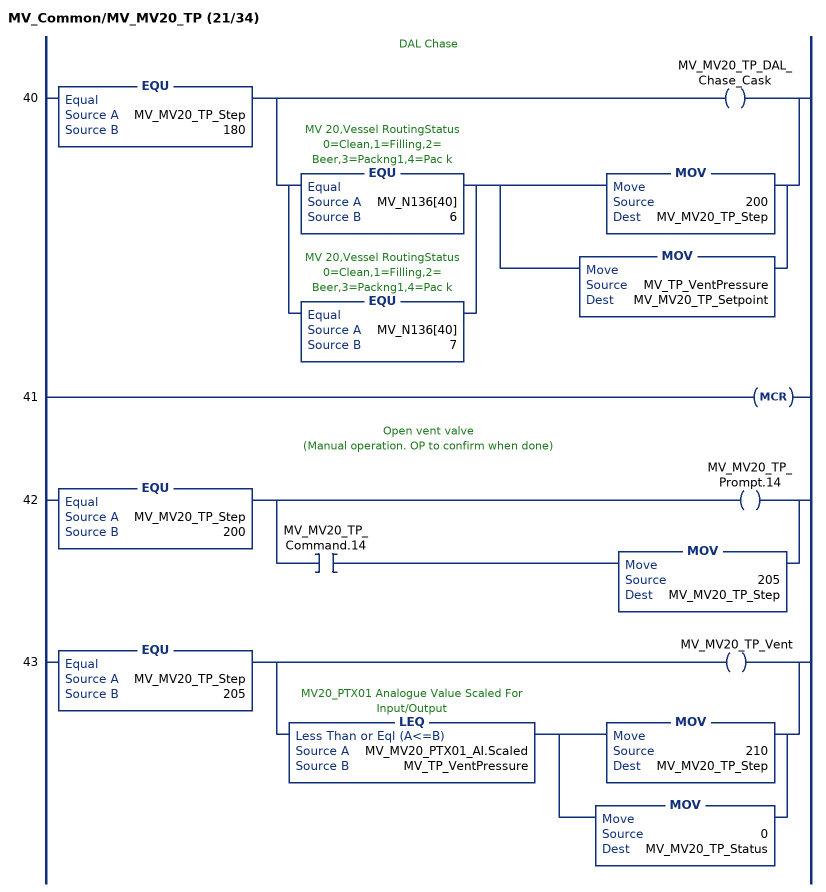
   // DAL Chase
   40: EQU(MV_MV20_TP_Step,180)[OTE(MV_MV20_TP_DAL_Chase_Cask) ,[EQU(MV_N136[40],6) ,EQU(MV_N136[40],7) ] [MOV(200,MV_MV20_TP_Step) ,MOV(MV_TP_VentPressure,MV_MV20_TP_Setpoint) ] ];
   41: MCR();
   // Open vent valve
   // (Manual operation. OP to confirm when done)
   42: EQU(MV_MV20_TP_Step,200)[OTE(MV_MV20_TP_Prompt.14) ,XIC(MV_MV20_TP_Command.14) MOV(205,MV_MV20_TP_Step) ];
   43: EQU(MV_MV20_TP_Step,205)[OTE(MV_MV20_TP_Vent) ,LEQ(MV_MV20_PTX01_AI.Scaled,MV_TP_VentPressure) [MOV(210,MV_MV20_TP_Step) ,MOV(0,MV_MV20_TP_Status) ] ];
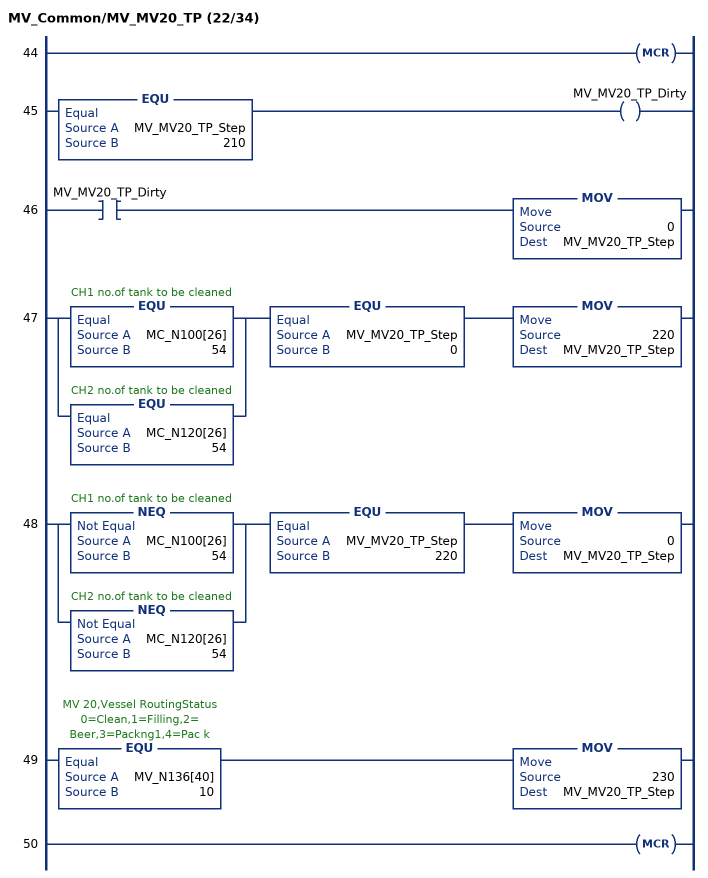
   44: MCR();
   45: EQU(MV_MV20_TP_Step,210)OTE(MV_MV20_TP_Dirty);
   46: XIC(MV_MV20_TP_Dirty)MOV(0,MV_MV20_TP_Step);
   47: [EQU(MC_N100[26],54) ,EQU(MC_N120[26],54) ]EQU(MV_MV20_TP_Step,0)MOV(220,MV_MV20_TP_Step);
   48: [NEQ(MC_N100[26],54) ,NEQ(MC_N120[26],54) ]EQU(MV_MV20_TP_Step,220)MOV(0,MV_MV20_TP_Step);
   49: EQU(MV_N136[40],10)MOV(230,MV_MV20_TP_Step);
   50: MCR();
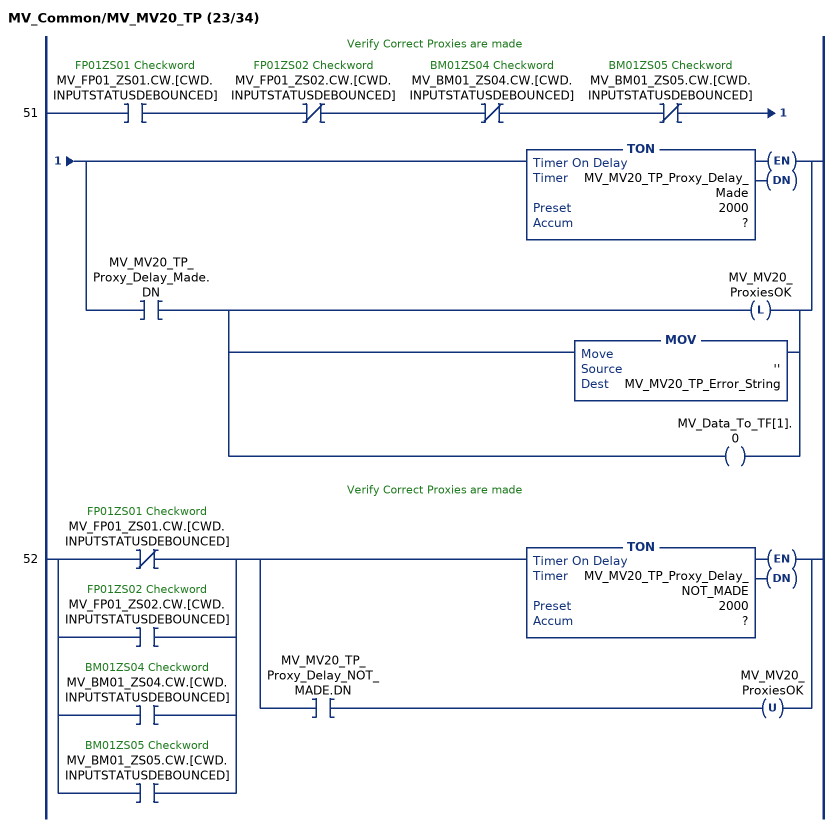
   // Verify Correct Proxies are made
   51: XIC(MV_FP01_ZS01.CW.[CWD.INPUTSTATUSDEBOUNCED])XIO(MV_FP01_ZS02.CW.[CWD.INPUTSTATUSDEBOUNCED])XIO(MV_BM01_ZS04.CW.[CWD.INPUTSTATUSDEBOUNCED])XIO(MV_BM01_ZS05.CW.[CWD.INPUTSTATUSDEBOUNCED])[TON(MV_MV20_TP_Proxy_Delay_Made,?,?) ,XIC(MV_MV20_TP_Proxy_Delay_Made.DN) [OTL(MV_MV20_ProxiesOK) ,MOV('',MV_MV20_TP_Error_String) ,OTE(MV_Data_To_TF[1].0) ] ];
   // Verify Correct Proxies are made
   52: [XIO(MV_FP01_ZS01.CW.[CWD.INPUTSTATUSDEBOUNCED]) ,XIC(MV_FP01_ZS02.CW.[CWD.INPUTSTATUSDEBOUNCED]) ,XIC(MV_BM01_ZS04.CW.[CWD.INPUTSTATUSDEBOUNCED]) ,XIC(MV_BM01_ZS05.CW.[CWD.INPUTSTATUSDEBOUNCED]) ][TON(MV_MV20_TP_Proxy_Delay_NOT_MADE,?,?) ,XIC(MV_MV20_TP_Proxy_Delay_NOT_MADE.DN) OTU(MV_MV20_ProxiesOK) ];
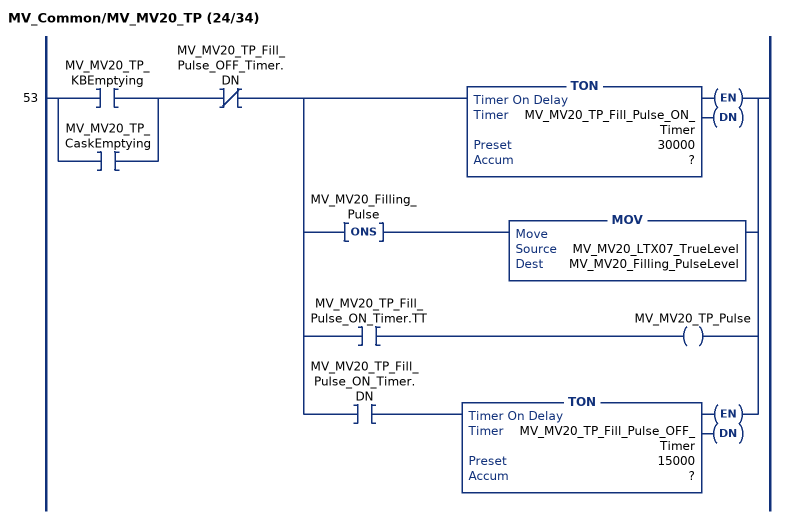
   53: [XIC(MV_MV20_TP_KBEmptying) ,XIC(MV_MV20_TP_CaskEmptying) ]XIO(MV_MV20_TP_Fill_Pulse_OFF_Timer.DN)[TON(MV_MV20_TP_Fill_Pulse_ON_Timer,?,?) ,ONS(MV_MV20_Filling_Pulse) MOV(MV_MV20_LTX07_TrueLevel,MV_MV20_Filling_PulseLevel) ,XIC(MV_MV20_TP_Fill_Pulse_ON_Timer.TT) OTE(MV_MV20_TP_Pulse) ,XIC(MV_MV20_TP_Fill_Pulse_ON_Timer.DN) TON(MV_MV20_TP_Fill_Pulse_OFF_Timer,?,?) ];
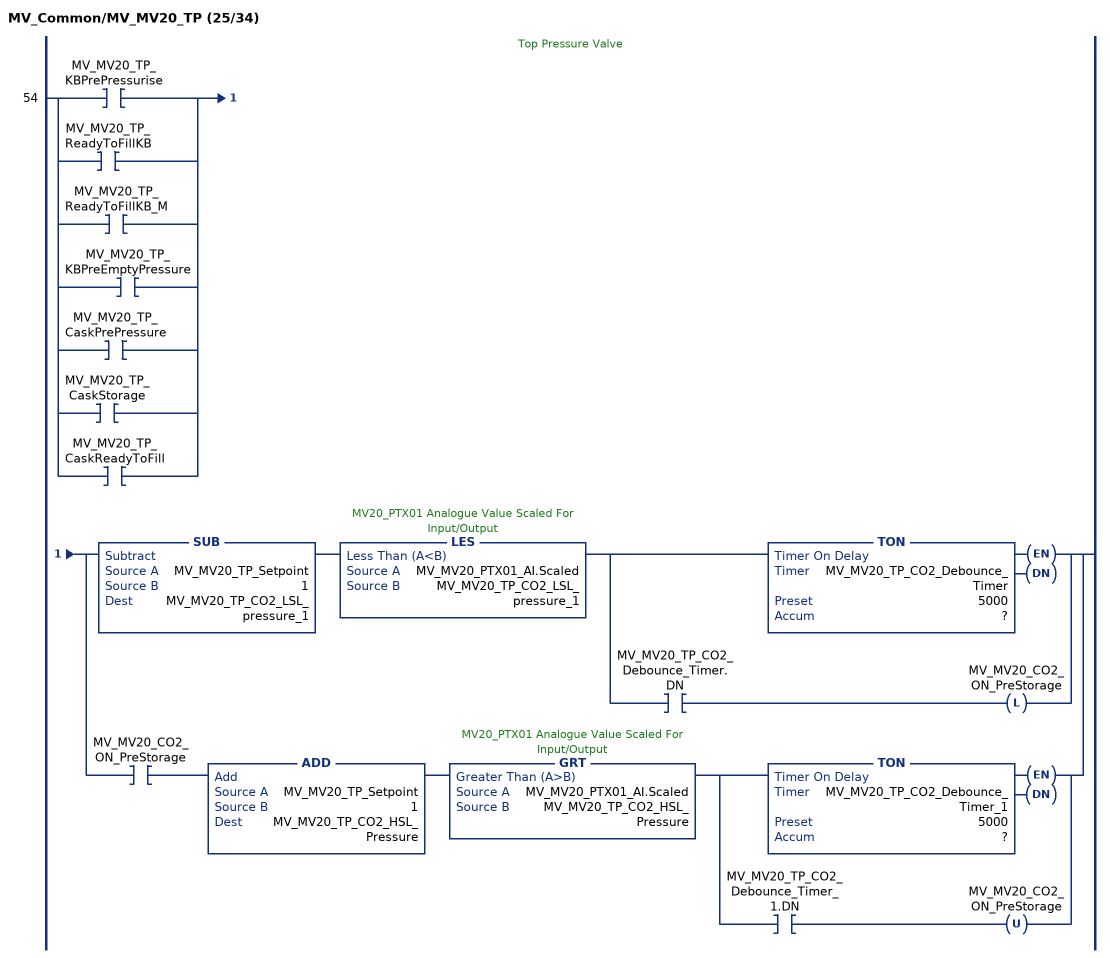
   // Top Pressure Valve
   54: [XIC(MV_MV20_TP_KBPrePressurise) ,XIC(MV_MV20_TP_ReadyToFillKB) ,XIC(MV_MV20_TP_ReadyToFillKB_M) ,XIC(MV_MV20_TP_KBPreEmptyPressure) ,XIC(MV_MV20_TP_CaskPrePressure) ,XIC(MV_MV20_TP_CaskStorage) ,XIC(MV_MV20_TP_CaskReadyToFill) ][SUB(MV_MV20_TP_Setpoint,1,MV_MV20_TP_CO2_LSL_pressure_1) LES(MV_MV20_PTX01_AI.Scaled,MV_MV20_TP_CO2_LSL_pressure_1) [TON(MV_MV20_TP_CO2_Debounce_Timer,?,?) ,XIC(MV_MV20_TP_CO2_Debounce_Timer.DN) OTL(MV_MV20_CO2_ON_PreStorage) ] ,XIC(MV_MV20_CO2_ON_PreStorage) ADD(MV_MV20_TP_Setpoint,1,MV_MV20_TP_CO2_HSL_Pressure) GRT(MV_MV20_PTX01_AI.Scaled,MV_MV20_TP_CO2_HSL_Pressure) [TON(MV_MV20_TP_CO2_Debounce_Timer_1,?,?) ,XIC(MV_MV20_TP_CO2_Debounce_Timer_1.DN) OTU(MV_MV20_CO2_ON_PreStorage) ] ];
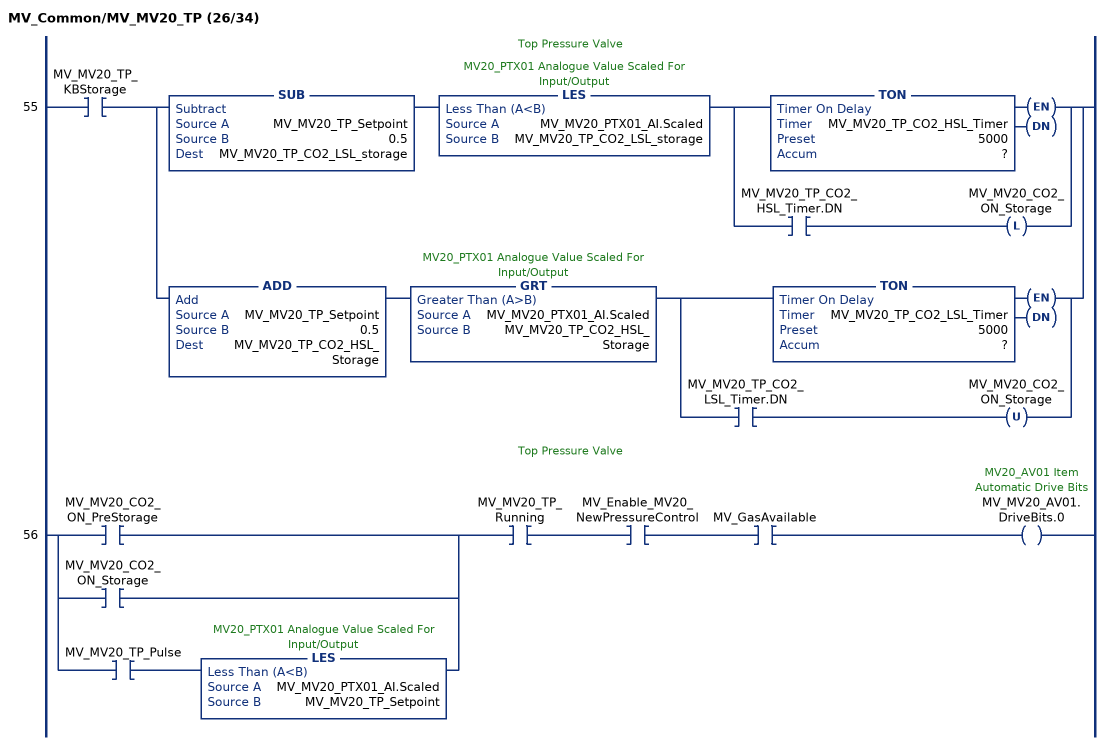
   // Top Pressure Valve
   55: XIC(MV_MV20_TP_KBStorage)[SUB(MV_MV20_TP_Setpoint,0.5,MV_MV20_TP_CO2_LSL_storage) LES(MV_MV20_PTX01_AI.Scaled,MV_MV20_TP_CO2_LSL_storage) [TON(MV_MV20_TP_CO2_HSL_Timer,?,?) ,XIC(MV_MV20_TP_CO2_HSL_Timer.DN) OTL(MV_MV20_CO2_ON_Storage) ] ,ADD(MV_MV20_TP_Setpoint,0.5,MV_MV20_TP_CO2_HSL_Storage) GRT(MV_MV20_PTX01_AI.Scaled,MV_MV20_TP_CO2_HSL_Storage) [TON(MV_MV20_TP_CO2_LSL_Timer,?,?) ,XIC(MV_MV20_TP_CO2_LSL_Timer.DN) OTU(MV_MV20_CO2_ON_Storage) ] ];
   // Top Pressure Valve
   56: [XIC(MV_MV20_CO2_ON_PreStorage) ,XIC(MV_MV20_CO2_ON_Storage) ,XIC(MV_MV20_TP_Pulse) LES(MV_MV20_PTX01_AI.Scaled,MV_MV20_TP_Setpoint) ]XIC(MV_MV20_TP_Running)XIC(MV_Enable_MV20_NewPressureControl)XIC(MV_GasAvailable)OTE(MV_MV20_AV01.DriveBits.0);
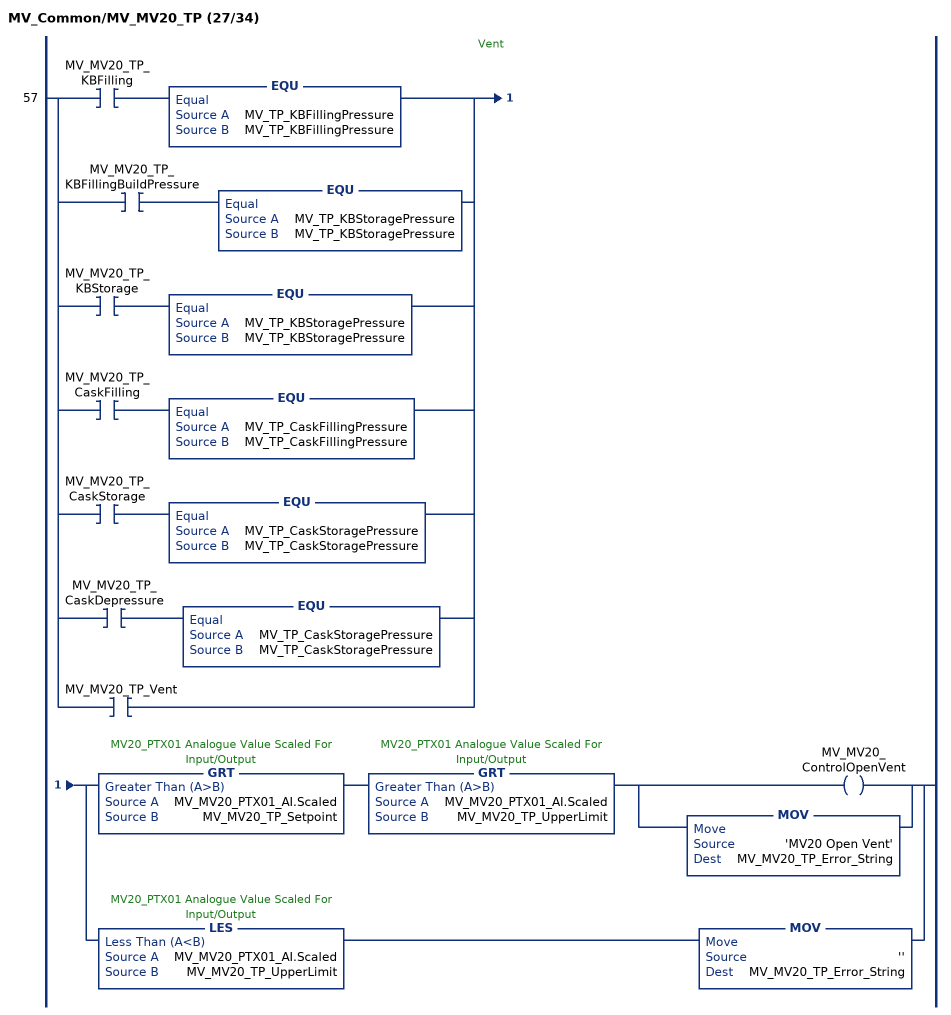
   // Vent
   57: [XIC(MV_MV20_TP_KBFilling) EQU(MV_TP_KBFillingPressure,MV_TP_KBFillingPressure) ,XIC(MV_MV20_TP_KBFillingBuildPressure) EQU(MV_TP_KBStoragePressure,MV_TP_KBStoragePressure) ,XIC(MV_MV20_TP_KBStorage) EQU(MV_TP_KBStoragePressure,MV_TP_KBStoragePressure) ,XIC(MV_MV20_TP_CaskFilling) EQU(MV_TP_CaskFillingPressure,MV_TP_CaskFillingPressure) ,XIC(MV_MV20_TP_CaskStorage) EQU(MV_TP_CaskStoragePressure,MV_TP_CaskStoragePressure) ,XIC(MV_MV20_TP_CaskDepressure) EQU(MV_TP_CaskStoragePressure,MV_TP_CaskStoragePressure) ,XIC(MV_MV20_TP_Vent) ][GRT(MV_MV20_PTX01_AI.Scaled,MV_MV20_TP_Setpoint) GRT(MV_MV20_PTX01_AI.Scaled,MV_MV20_TP_UpperLimit) [OTE(MV_MV20_ControlOpenVent) ,MOV('MV20 Open Vent',MV_MV20_TP_Error_String) ] ,LES(MV_MV20_PTX01_AI.Scaled,MV_MV20_TP_UpperLimit) MOV('',MV_MV20_TP_Error_String) ];
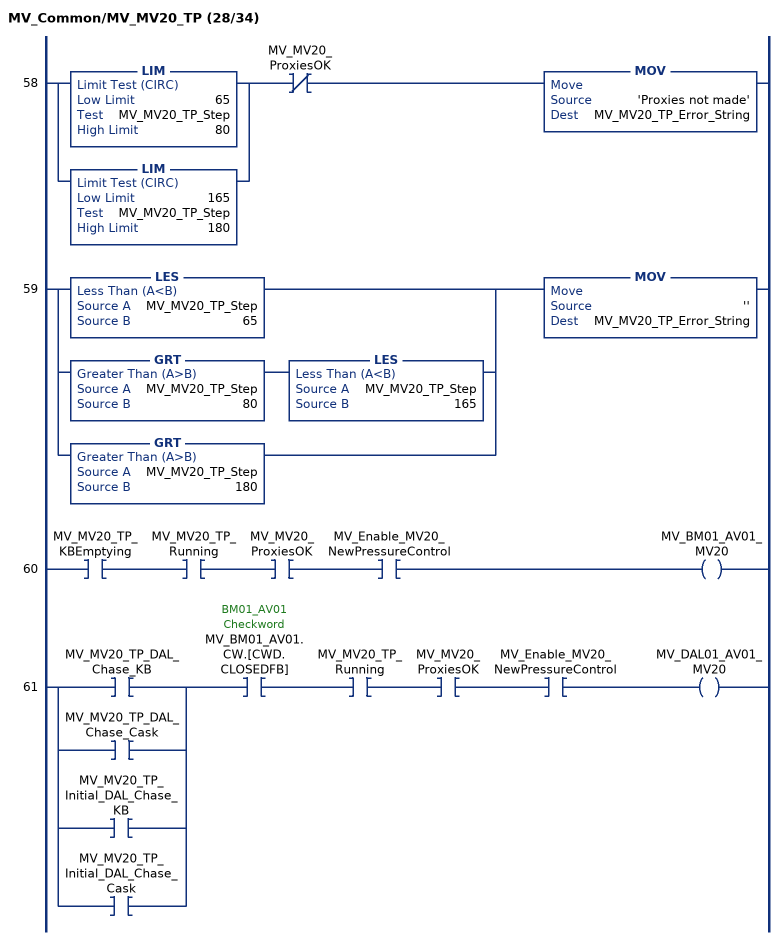
   58: [LIM(65,MV_MV20_TP_Step,80) ,LIM(165,MV_MV20_TP_Step,180) ]XIO(MV_MV20_ProxiesOK)MOV('Proxies not made',MV_MV20_TP_Error_String);
   59: [LES(MV_MV20_TP_Step,65) ,GRT(MV_MV20_TP_Step,80) LES(MV_MV20_TP_Step,165) ,GRT(MV_MV20_TP_Step,180) ]MOV('',MV_MV20_TP_Error_String);
   60: XIC(MV_MV20_TP_KBEmptying)XIC(MV_MV20_TP_Running)XIC(MV_MV20_ProxiesOK)XIC(MV_Enable_MV20_NewPressureControl)OTE(MV_BM01_AV01_MV20);
   61: [XIC(MV_MV20_TP_DAL_Chase_KB) ,XIC(MV_MV20_TP_DAL_Chase_Cask) ,XIC(MV_MV20_TP_Initial_DAL_Chase_KB) ,XIC(MV_MV20_TP_Initial_DAL_Chase_Cask) ]XIC(MV_BM01_AV01.CW.[CWD.CLOSEDFB])XIC(MV_MV20_TP_Running)XIC(MV_MV20_ProxiesOK)XIC(MV_Enable_MV20_NewPressureControl)OTE(MV_DAL01_AV01_MV20);
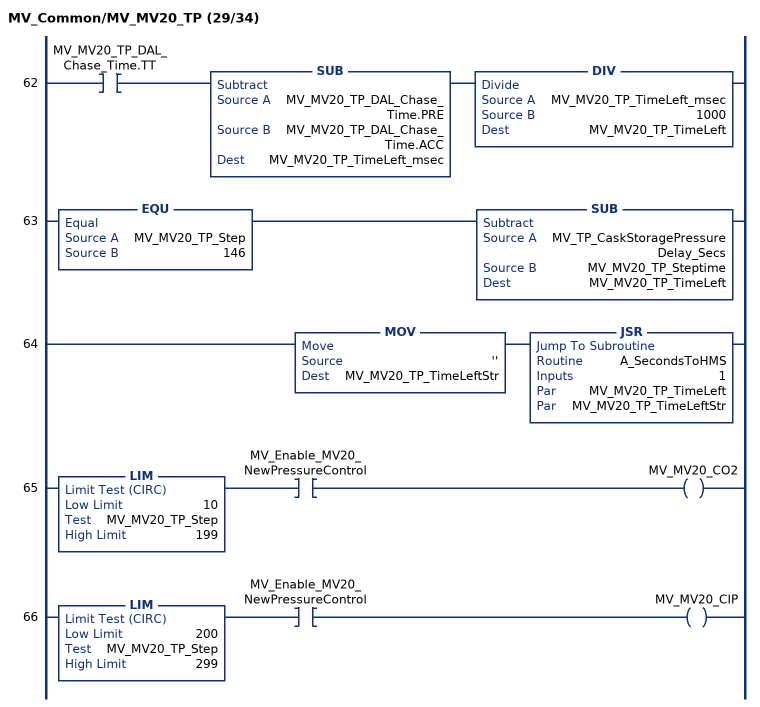
   62: XIC(MV_MV20_TP_DAL_Chase_Time.TT)SUB(MV_MV20_TP_DAL_Chase_Time.PRE,MV_MV20_TP_DAL_Chase_Time.ACC,MV_MV20_TP_TimeLeft_msec)DIV(MV_MV20_TP_TimeLeft_msec,1000,MV_MV20_TP_TimeLeft);
   63: EQU(MV_MV20_TP_Step,146)SUB(MV_TP_CaskStoragePressureDelay_Secs,MV_MV20_TP_Steptime,MV_MV20_TP_TimeLeft);
   64: MOV('',MV_MV20_TP_TimeLeftStr)JSR(A_SecondsToHMS,1,MV_MV20_TP_TimeLeft,MV_MV20_TP_TimeLeftStr);
   65: LIM(10,MV_MV20_TP_Step,199)XIC(MV_Enable_MV20_NewPressureControl)OTE(MV_MV20_CO2);
   66: LIM(200,MV_MV20_TP_Step,299)XIC(MV_Enable_MV20_NewPressureControl)OTE(MV_MV20_CIP);
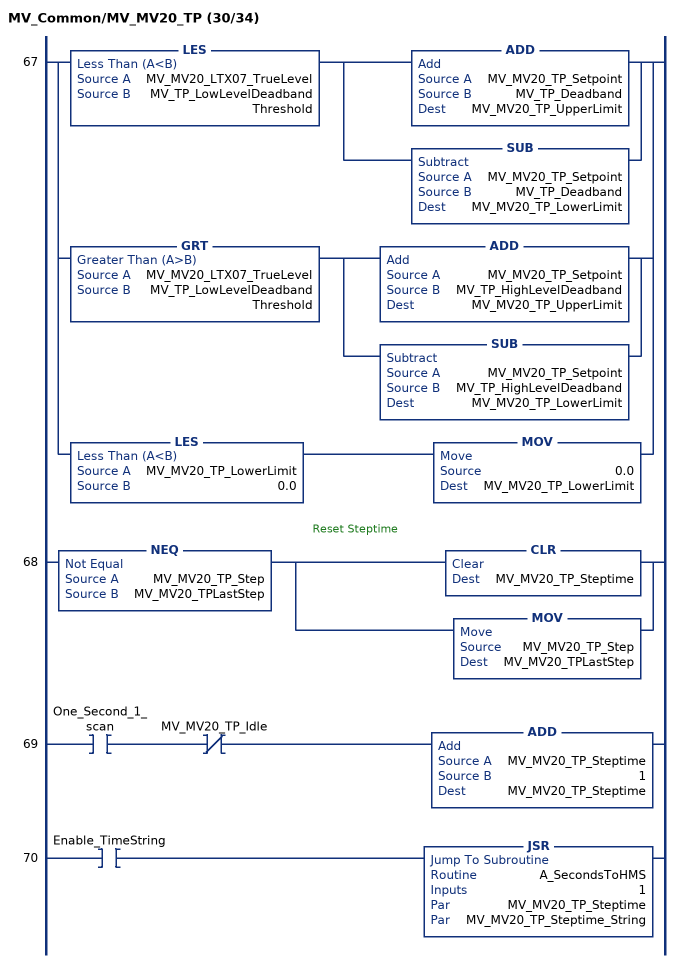
   67: [LES(MV_MV20_LTX07_TrueLevel,MV_TP_LowLevelDeadbandThreshold) [ADD(MV_MV20_TP_Setpoint,MV_TP_Deadband,MV_MV20_TP_UpperLimit) ,SUB(MV_MV20_TP_Setpoint,MV_TP_Deadband,MV_MV20_TP_LowerLimit) ] ,GRT(MV_MV20_LTX07_TrueLevel,MV_TP_LowLevelDeadbandThreshold) [ADD(MV_MV20_TP_Setpoint,MV_TP_HighLevelDeadband,MV_MV20_TP_UpperLimit) ,SUB(MV_MV20_TP_Setpoint,MV_TP_HighLevelDeadband,MV_MV20_TP_LowerLimit) ] ,LES(MV_MV20_TP_LowerLimit,0.0) MOV(0.0,MV_MV20_TP_LowerLimit) ];
   // Reset Steptime
   68: NEQ(MV_MV20_TP_Step,MV_MV20_TPLastStep)[CLR(MV_MV20_TP_Steptime) ,MOV(MV_MV20_TP_Step,MV_MV20_TPLastStep) ];
   69: XIC(One_Second_1_scan)XIO(MV_MV20_TP_Idle)ADD(MV_MV20_TP_Steptime,1,MV_MV20_TP_Steptime);
   70: XIC(Enable_TimeString)JSR(A_SecondsToHMS,1,MV_MV20_TP_Steptime,MV_MV20_TP_Steptime_String);
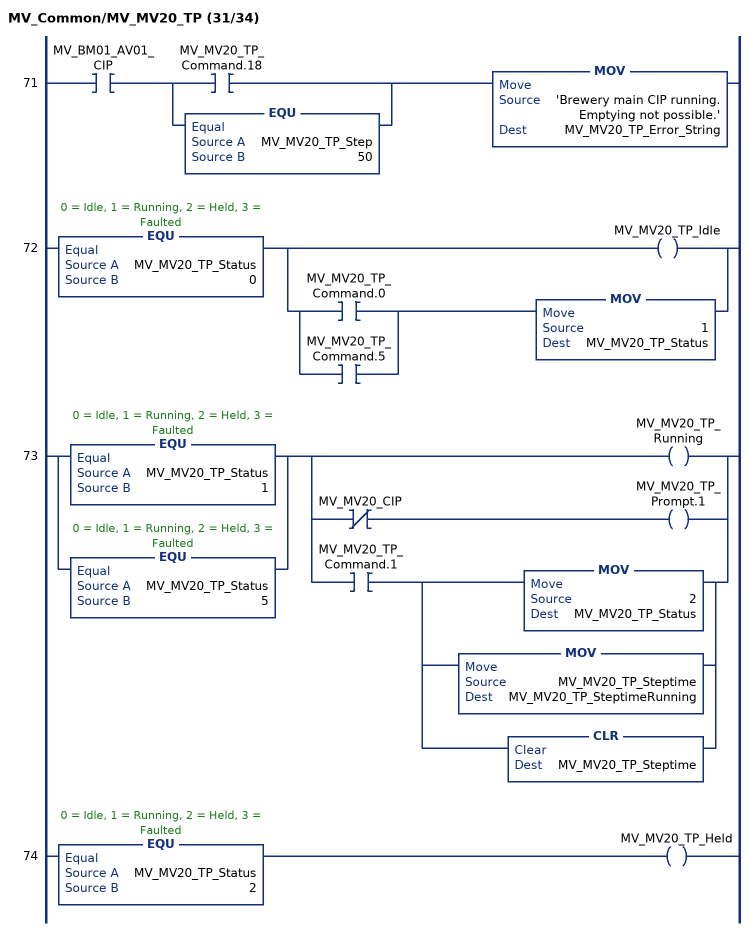
   71: XIC(MV_BM01_AV01_CIP)[XIC(MV_MV20_TP_Command.18) ,EQU(MV_MV20_TP_Step,50) ]MOV('Brewery main CIP running. Emptying not possible.',MV_MV20_TP_Error_String);
   72: EQU(MV_MV20_TP_Status,0)[OTE(MV_MV20_TP_Idle) ,[XIC(MV_MV20_TP_Command.0) ,XIC(MV_MV20_TP_Command.5) ] MOV(1,MV_MV20_TP_Status) ];
   73: [EQU(MV_MV20_TP_Status,1) ,EQU(MV_MV20_TP_Status,5) ][OTE(MV_MV20_TP_Running) ,XIO(MV_MV20_CIP) OTE(MV_MV20_TP_Prompt.1) ,XIC(MV_MV20_TP_Command.1) [MOV(2,MV_MV20_TP_Status) ,MOV(MV_MV20_TP_Steptime,MV_MV20_TP_SteptimeRunning) ,CLR(MV_MV20_TP_Steptime) ] ];
   74: EQU(MV_MV20_TP_Status,2)OTE(MV_MV20_TP_Held);
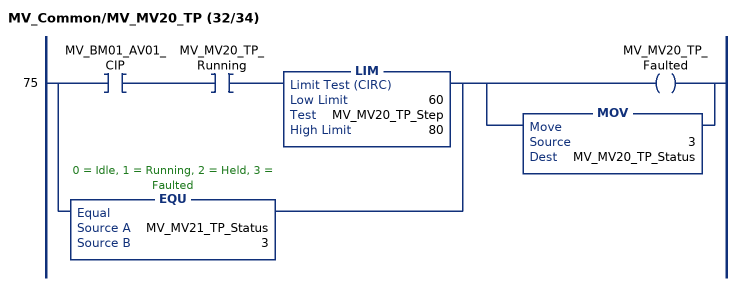
   75: [XIC(MV_BM01_AV01_CIP) XIC(MV_MV20_TP_Running) LIM(60,MV_MV20_TP_Step,80) ,EQU(MV_MV21_TP_Status,3) ][OTE(MV_MV20_TP_Faulted) ,MOV(3,MV_MV20_TP_Status) ];
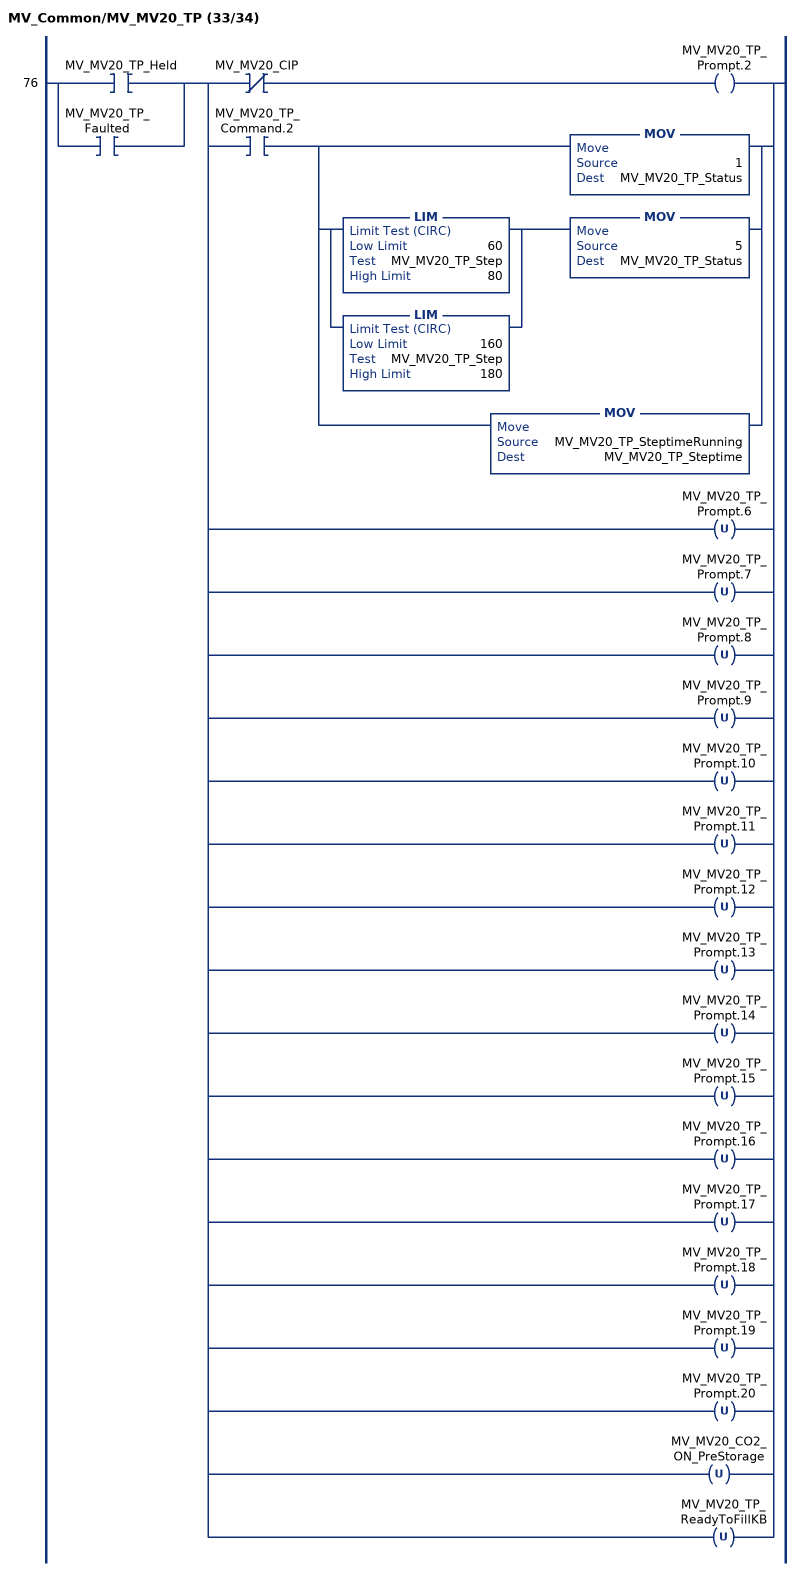
   76: [XIC(MV_MV20_TP_Held) ,XIC(MV_MV20_TP_Faulted) ][XIO(MV_MV20_CIP) OTE(MV_MV20_TP_Prompt.2) ,XIC(MV_MV20_TP_Command.2) [MOV(1,MV_MV20_TP_Status) ,[LIM(60,MV_MV20_TP_Step,80) ,LIM(160,MV_MV20_TP_Step,180) ] MOV(5,MV_MV20_TP_Status) ,MOV(MV_MV20_TP_SteptimeRunning,MV_MV20_TP_Steptime) ] ,OTU(MV_MV20_TP_Prompt.6) ,OTU(MV_MV20_TP_Prompt.7) ,OTU(MV_MV20_TP_Prompt.8) ,OTU(MV_MV20_TP_Prompt.9) ,OTU(MV_MV20_TP_Prompt.10) ,OTU(MV_MV20_TP_Prompt.11) ,OTU(MV_MV20_TP_Prompt.12) ,OTU(MV_MV20_TP_Prompt.13) ,OTU(MV_MV20_TP_Prompt.14) ,OTU(MV_MV20_TP_Prompt.15) ,OTU(MV_MV20_TP_Prompt.16) ,OTU(MV_MV20_TP_Prompt.17) ,OTU(MV_MV20_TP_Prompt.18) ,OTU(MV_MV20_TP_Prompt.19) ,OTU(MV_MV20_TP_Prompt.20) ,OTU(MV_MV20_CO2_ON_PreStorage) ,OTU(MV_MV20_TP_ReadyToFillKB) ];
